
           REGION "GET ARRAY PARAMETERS"
               #len.tblData := UDINT_TO_DINT(CountOfElements(#tblData));
               #len.tblDisp := UDINT_TO_DINT(CountOfElements(#tblDisp));
           END_REGION

           REGION "CALCULATE UPPER BOUND"
               #ubound := #len.tblData;
               IF #first_null_index <= #len.tblData THEN
                   IF #first_null_index > 0 THEN
                       #ubound := #first_null_index;
                   END_IF;
               END_IF;
           END_REGION


           REGION "CALCULATE OFFSET"
               #offset := "Table Nav: Calculate Offset"(pulses := #pulses,
                                                        lenTblData := #ubound,
                                                        lenTblDisp := #len.tblDisp,
                                                        r1 := #r1);
           END_REGION


           REGION "CALCULATE FIRST ROW"
               #r1 := "Table Nav: Get First Row"(table_length := #ubound,
                                                 offset := #offset,
                                                 first_row := #r1);
           END_REGION


           REGION "CALCUALTE ROW INDICIES"
               "Table Nav: Calc Row Indices"(lenTblData := #ubound,
                                             lenTblDisp := #len.tblDisp,
                                             r1 := #r1,
                                             rowIndicies := #ret_row_indices);
           END_REGION


           REGION "RETURN ROW INDICIES"
               #RET_VAL := MOVE_BLK_VARIANT(SRC := #ret_row_indices,
                                            COUNT := DINT_TO_UDINT(#len.tblDisp),
                                            SRC_INDEX := 0,
                                            DEST_INDEX := 0,
                                            DEST => #rowIndices);
           END_REGION

       END_IF;
   END_REGION
END_FUNCTION_BLOCK

FUNCTION_BLOCK "Table Nav: Pulses"   // FB44, SCL
{ S7_Optimized_Access := 'TRUE' }
VERSION : 0.1
   VAR_INPUT
      press : "Nav Bar Data: PLC";
   END_VAR
   VAR_OUTPUT
      pulses : "Nav Bar Data: PLC";
   END_VAR
   VAR
      old : "Nav Bar Data: PLC";
   END_VAR
BEGIN
   REGION "EVALUATION"
       #pulses.top.actuate := #press.top.actuate AND NOT #old.top.actuate;
       #pulses.pageUp.actuate := #press.pageUp.actuate AND NOT #old.pageUp.actuate;
       #pulses.lineUp.actuate := #press.lineUp.actuate AND NOT #old.lineUp.actuate;
       #pulses.lineDown.actuate := #press.lineDown.actuate AND NOT #old.lineDown.actuate;
       #pulses.pageDown.actuate := #press.pageDown.actuate AND NOT #old.pageDown.actuate;
       #pulses.bottom.actuate := #press.bottom.actuate AND NOT #old.bottom.actuate;
   END_REGION

   REGION "CHANGE DETECTION"
       #old.top.actuate := #press.top.actuate;
       #old.pageUp.actuate := #press.pageUp.actuate;
       #old.lineUp.actuate := #press.lineUp.actuate;
       #old.lineDown.actuate := #press.lineDown.actuate;
       #old.pageDown.actuate := #press.pageDown.actuate;
       #old.bottom.actuate := #press.bottom.actuate;
   END_REGION
END_FUNCTION_BLOCK

FUNCTION "Table Nav: Get Null Index" : DInt   // FC14, SCL
{ S7_Optimized_Access := 'TRUE' }
VERSION : 0.1
   VAR_INPUT
      nullFlag : Int;
      nullCheckVals : Array[0.."WIP_COUNT"] of DInt;
   END_VAR
   VAR_TEMP
      pNullCheck : DInt;
   END_VAR
BEGIN
   WHILE #nullCheckVals[#pNullCheck] <> #nullFlag AND #pNullCheck <= "WIP_COUNT" DO
       #pNullCheck += 1;
   END_WHILE;
   #"Table Nav: Get Null Index" := #pNullCheck;
END_FUNCTION

FUNCTION "Table Nav: Get First Row" : DInt   // FC44, SCL
{ S7_Optimized_Access := 'TRUE' }
VERSION : 0.1
   VAR_INPUT
      first_row : DInt;
      offset : DInt;
      table_length : DInt;
   END_VAR
   VAR_TEMP
      ret : DInt;
   END_VAR
BEGIN
   REGION "DESCRIPTION"
       (*
       The new first row of the table is calculated from the offset. 
       Rollover and rollunder are resolved for the first row.
       *)
   END_REGION

   REGION "COPY TO INTERNAL"
       #ret := #first_row + #offset;
   END_REGION

   REGION "ROLLUNDER"
       IF #ret < 0 THEN
           #ret := #ret + #table_length;
       END_IF;
   END_REGION

   REGION "ROLLOVER"
       IF #ret > #table_length THEN
           #ret := #ret - #table_length;
       END_IF;
   END_REGION

   REGION "OUTPUT"
       #"Table Nav: Get First Row" := #ret;
   END_REGION
END_FUNCTION

FUNCTION "Table Nav: Calculate Offset" : DInt   // FC45, SCL
{ S7_Optimized_Access := 'TRUE' }
VERSION : 0.1
   VAR_INPUT
      lenTblData : DInt;
      lenTblDisp : DInt;
      pulses : "Nav Bar Data: PLC";
      r1 : DInt;
   END_VAR
   VAR_TEMP
      retOffset : DInt;
   END_VAR
   // Ret_Val : offset from table row 1 from button
BEGIN
   REGION "DESCRIPTION"
       (*
       The offset from the first row of the table is calculated based on the button pressed.
       *)
   END_REGION

   REGION "TOP"
       IF #pulses.top.actuate THEN
           #retOffset := -1 * #r1;
       END_IF;
   END_REGION

   REGION "PAGE UP"
       IF #pulses.pageUp.actuate THEN
           #retOffset := -1 * #lenTblDisp;
       END_IF;
   END_REGION

   REGION "LINE UP"
       IF #pulses.lineUp.actuate THEN
           #retOffset := -1;
       END_IF;
   END_REGION

   REGION "LINE DOWN"
       IF #pulses.lineDown.actuate THEN
           #retOffset := 1;
       END_IF;
   END_REGION

   REGION "PAGE DOWN"
       IF #pulses.pageDown.actuate THEN
           #retOffset := #lenTblDisp ;
       END_IF;
   END_REGION

   REGION "BOTTOM"
       IF #pulses.bottom.actuate THEN
           #retOffset := #lenTblData - #lenTblDisp - #r1;
       END_IF;
   END_REGION

   REGION "RETURN"
       #"Table Nav: Calculate Offset" := #retOffset;
   END_REGION
END_FUNCTION

FUNCTION "Table Nav: Calc Row Indices" : Void   // FC46, SCL
{ S7_Optimized_Access := 'TRUE' }
VERSION : 0.1
   VAR_INPUT
      lenTblData : DInt;
      lenTblDisp : DInt;
      r1 : DInt;
   END_VAR
   VAR_IN_OUT
      rowIndicies : Array[0..#lenRetArr] of DInt;
   END_VAR
   VAR_TEMP
      pOutArr : Int;
      calcRowIdx : DInt;
      retRowIndicies : Array[0..#lenRetArr] of DInt;
   END_VAR
   VAR CONSTANT
      lenRetArr : Int := 999;
   END_VAR
BEGIN
   REGION "DESCRIPTION"
       (*
       An array of the row indicies that the table should display is returned.
       Rollover and rollunder are calculated index by index.
       *) 
   END_REGION

   REGION "INITIALIZE OUTPUT"
       FOR #pOutArr := 0 TO #lenRetArr DO
           #rowIndicies[#pOutArr] := 0;
       END_FOR;
   END_REGION

   REGION "CALCULATE INDICIES"
       FOR #pOutArr := 0 TO DINT_TO_INT(#lenTblDisp) DO

           REGION "CALCULATE INDEX"
               #calcRowIdx := #r1 + INT_TO_DINT(#pOutArr);
           END_REGION

           REGION "ROLL UNDER"
               IF #calcRowIdx < 0 THEN
                   #calcRowIdx := #calcRowIdx + #lenTblDisp;
               END_IF;
           END_REGION

           REGION "ROLL OVER"
               IF #calcRowIdx >= #lenTblData THEN
                   #calcRowIdx := #calcRowIdx - #lenTblData;
               END_IF;
           END_REGION

           REGION "SAVE TO ARRAY"
               #retRowIndicies[#pOutArr] := #calcRowIdx;
           END_REGION

       END_FOR;
   END_REGION

   REGION "OUTPUT"
       #rowIndicies := #retRowIndicies;
   END_REGION
END_FUNCTION

FUNCTION "Table Nav: Run Trigger" : Bool   // FC47, SCL
{ S7_Optimized_Access := 'TRUE' }
VERSION : 0.1
   VAR_INPUT
      pulses : "Nav Bar Data: PLC";
   END_VAR
BEGIN
   #"Table Nav: Run Trigger" :=
       #pulses.top.actuate OR
       #pulses.pageUp.actuate OR
       #pulses.lineUp.actuate OR
       #pulses.lineDown.actuate OR
       #pulses.pageDown.actuate OR
       #pulses.bottom.actuate;
END_FUNCTION

// folder: Utilities/Time

FUNCTION "Time.to_WString" : WString   // FC36, SCL
{ S7_Optimized_Access := 'TRUE' }
VERSION : 0.1
   VAR_INPUT
      "Time" : Time;
   END_VAR
   VAR_TEMP
      _time : DInt;
      _days : DInt;
      _hours : DInt;
      _minutes : DInt;
      _seconds : DInt;
      "Time Elements" : Array[0..4] of WString;
      Length : Int;
      _return : WString;
   END_VAR
   VAR CONSTANT
      COLON : WString := WSTRING#':';
   END_VAR
BEGIN
   REGION GET INPUT
       #_time := #Time;
   END_REGION


   REGION CONVERT TIME INTO INDIVIDUAL PLACE VALUES
       #_days := "Time.Get_Days"(#_time);
       #_hours := "Time.Get_MOD_Hours"(#_time);
       #_minutes := "Time.Get_MOD_Minutes"(#_time);
       #_seconds := "Time.Get_MOD_Seconds"(#_time);
   END_REGION


   REGION "ASSEMBLE DISPLAY STRING"
       IF #_days > 0 THEN
           #_return := CONCAT_WSTRING(IN1 := #_return, IN2 := "Time.to_WString.Days"(#_time), IN3 := #COLON);
           #_return := CONCAT_WSTRING(IN1 := #_return, IN2 := "Time.to_WString.MOD_Hours"(#_time), IN3 := #COLON);
           #_return := CONCAT_WSTRING(IN1 := #_return, IN2 := "Time.to_WString.MOD_Minutes"(#_time), IN3 := #COLON);
           #_return := CONCAT_WSTRING(IN1 := #_return, IN2 := "Time.to_WString.MOD_Seconds"(#_time));
           #"Time.to_WString" := #_return;
           RETURN;
       END_IF;
       IF #_hours > 0 THEN
           #_return := CONCAT_WSTRING(IN1 := #_return, IN2 := "Time.to_WString.MOD_Hours"(#_time), IN3 := #COLON);
           #_return := CONCAT_WSTRING(IN1 := #_return, IN2 := "Time.to_WString.MOD_Minutes"(#_time), IN3 := #COLON);
           #_return := CONCAT_WSTRING(IN1 := #_return, IN2 := "Time.to_WString.MOD_Seconds"(#_time));
           #"Time.to_WString" := #_return;
           RETURN;
       END_IF;
       IF #_minutes > 0 THEN
           #_return := CONCAT_WSTRING(IN1 := #_return, IN2 := "Time.to_WString.MOD_Minutes"(#_time), IN3 := #COLON);
           #_return := CONCAT_WSTRING(IN1 := #_return, IN2 := "Time.to_WString.MOD_Seconds"(#_time));
           #"Time.to_WString" := #_return;
           RETURN;
       END_IF;
       IF #_seconds > 0 THEN
           #_return := CONCAT_WSTRING(IN1 := #_return, IN2 := "Time.to_WString.MOD_Seconds"(#_time));
           #"Time.to_WString" := #_return;
           RETURN;
       END_IF;
       #_return := WSTRING#'00:00';
       #"Time.to_WString" := #_return;
       RETURN;
   END_REGION
END_FUNCTION

FUNCTION "Time.to_WString.Seconds" : WString   // FC275, SCL
{ S7_Optimized_Access := 'TRUE' }
VERSION : 0.1
   VAR_INPUT
      value : Time;
   END_VAR
BEGIN
   #"Time.to_WString.Seconds" := "Time.to_WString.Prepare_Component"("Time.Get_Seconds"(#value));
END_FUNCTION

FUNCTION "Time.Get_MOD_Seconds" : DInt   // FC276, SCL
{ S7_Optimized_Access := 'TRUE' }
VERSION : 0.1
   VAR_INPUT
      value : Time;
   END_VAR
   VAR CONSTANT
      SECONDS_PER_MINUTE : DInt := 60;
   END_VAR
BEGIN
   #"Time.Get_MOD_Seconds" := "Time.Get_Seconds"(#value) MOD #SECONDS_PER_MINUTE;
END_FUNCTION

FUNCTION "Time.Get_MOD_Minutes" : DInt   // FC277, SCL
{ S7_Optimized_Access := 'TRUE' }
VERSION : 0.1
   VAR_INPUT
      value : Time;
   END_VAR
   VAR CONSTANT
      MINUTES_PER_HOUR : DInt := 60;
   END_VAR
BEGIN
   #"Time.Get_MOD_Minutes" := "Time.Get_Minutes"(#value) MOD #MINUTES_PER_HOUR;
END_FUNCTION

FUNCTION "Time.Get_MOD_Hours" : DInt   // FC278, SCL
{ S7_Optimized_Access := 'TRUE' }
VERSION : 0.1
   VAR_INPUT
      value : Time;
   END_VAR
   VAR CONSTANT
      HOURS_PER_DAY : DInt := 24;
   END_VAR
BEGIN
   #"Time.Get_MOD_Hours" := "Time.Get_Hours"(#value) MOD #HOURS_PER_DAY;
END_FUNCTION

FUNCTION "Time.Get_Days" : Int   // FC279, SCL
{ S7_Optimized_Access := 'TRUE' }
VERSION : 0.1
   VAR_INPUT
      value : Time;
   END_VAR
   VAR_TEMP
      _return : DInt;
   END_VAR
   VAR CONSTANT
      MILLISECONDS_PER_DAY : DInt := 86_000_000;
   END_VAR
BEGIN
   #_return := #value / #MILLISECONDS_PER_DAY;
   #"Time.Get_Days" := DINT_TO_INT(#_return);
END_FUNCTION

FUNCTION "Time.Get_Seconds" : DInt   // FC280, SCL
{ S7_Optimized_Access := 'TRUE' }
VERSION : 0.1
   VAR_INPUT
      value : Time;
   END_VAR
   VAR CONSTANT
      MILLISECONDS_PER_SECOND : DInt := 1_000;
   END_VAR
BEGIN
   #"Time.Get_Seconds" := #value / #MILLISECONDS_PER_SECOND;
END_FUNCTION

FUNCTION "Time.Get_Minutes" : DInt   // FC281, SCL
{ S7_Optimized_Access := 'TRUE' }
VERSION : 0.1
   VAR_INPUT
      value : Time;
   END_VAR
   VAR CONSTANT
      MILLISECONDS_PER_MINUTE : DInt := 60_000;
   END_VAR
BEGIN
   #"Time.Get_Minutes" := #value / #MILLISECONDS_PER_MINUTE;
END_FUNCTION

FUNCTION "Time.to_WString.Prepare_Component" : WString   // FC282, SCL
{ S7_Optimized_Access := 'TRUE' }
VERSION : 0.1
   VAR_INPUT
      component : DInt;
   END_VAR
   VAR_TEMP
      _return : WString;
   END_VAR
   VAR CONSTANT
      ZERO : WChar := WCHAR#'0';
   END_VAR
BEGIN
   #_return := DINT_TO_WSTRING(#component);
   #_return := "Trim"("Strip Sign"(#_return));
   #_return := "Add Leading"("Leading Character" := #ZERO,
                             "Desired Length" := 2,
                             "String" := #_return);
   #"Time.to_WString.Prepare_Component" := #_return;
END_FUNCTION

FUNCTION "Time.to_WString.Minutes" : WString   // FC284, SCL
{ S7_Optimized_Access := 'TRUE' }
VERSION : 0.1
   VAR_INPUT
      value : Time;
   END_VAR
   VAR_TEMP
      _to_udint : UDInt;
      _return : WString;
   END_VAR
BEGIN
   #"Time.to_WString.Minutes" := "Time.to_WString.Prepare_Component"("Time.Get_Minutes"(#value));
END_FUNCTION

FUNCTION "Time.to_WString.MOD_Minutes" : WString   // FC285, SCL
{ S7_Optimized_Access := 'TRUE' }
VERSION : 0.1
   VAR_INPUT
      value : Time;
   END_VAR
BEGIN
   #"Time.to_WString.MOD_Minutes" := "Time.to_WString.Prepare_Component"("Time.Get_MOD_Minutes"(#value));
END_FUNCTION

FUNCTION "Time.to_WString.Hours" : WString   // FC286, SCL
{ S7_Optimized_Access := 'TRUE' }
VERSION : 0.1
   VAR_INPUT
      value : Time;
   END_VAR
BEGIN
   #"Time.to_WString.Hours" := "Time.to_WString.Prepare_Component"("Time.Get_Hours"(#value));
END_FUNCTION

FUNCTION "Time.to_WString.MOD_Seconds" : WString   // FC287, SCL
{ S7_Optimized_Access := 'TRUE' }
VERSION : 0.1
   VAR_INPUT
      value : Time;
   END_VAR
BEGIN
   #"Time.to_WString.MOD_Seconds" := "Time.to_WString.Prepare_Component"("Time.Get_MOD_Seconds"(#value));
END_FUNCTION

FUNCTION "Time.Get_Hours" : DInt   // FC288, SCL
{ S7_Optimized_Access := 'TRUE' }
VERSION : 0.1
   VAR_INPUT
      value : Time;
   END_VAR
   VAR CONSTANT
      MILLISECONDS_PER_HOUR : DInt := 3_600_000;
   END_VAR
BEGIN
   #"Time.Get_Hours" := #value / #MILLISECONDS_PER_HOUR;
END_FUNCTION

FUNCTION "Time.to_WString.MOD_Hours" : WString   // FC290, SCL
{ S7_Optimized_Access := 'TRUE' }
VERSION : 0.1
   VAR_INPUT
      value : Time;
   END_VAR
BEGIN
   #"Time.to_WString.MOD_Hours" := "Time.to_WString.Prepare_Component"("Time.Get_MOD_Hours"(#value));
END_FUNCTION

FUNCTION "Time.to_WString.Days" : WString   // FC291, SCL
{ S7_Optimized_Access := 'TRUE' }
VERSION : 0.1
   VAR_INPUT
      value : Time;
   END_VAR
BEGIN
   #"Time.to_WString.Days" := "Time.to_WString.Prepare_Component"("Time.Get_Days"(#value));
END_FUNCTION

// folder: Utilities/Timer

FUNCTION "Timer.WString_to_Real" : Real   // FC39, SCL
{ S7_Optimized_Access := 'TRUE' }
VERSION : 0.1
   VAR_INPUT
      wstring : WString;
   END_VAR
   VAR CONSTANT
      msPerSec : Real := 1000.0;
   END_VAR
BEGIN
   #"Timer.WString_to_Real" := DINT_TO_REAL(TIME_TO_DINT("WString.to_Time"(#wstring))) / #msPerSec;
END_FUNCTION

FUNCTION "Timer.Real_to_WString" : WString   // FC40, SCL
{ S7_Optimized_Access := 'TRUE' }
VERSION : 0.1
   VAR_INPUT
      realVal : Real;
   END_VAR
   VAR CONSTANT
      msPerSec : Real := 1000.0;
   END_VAR
BEGIN
   #"Timer.Real_to_WString" := "Time.to_WString"(DINT_TO_TIME(REAL_TO_DINT(#realVal * #msPerSec)));
END_FUNCTION

FUNCTION "Timer" : Void   // FC79, SCL
{ S7_Optimized_Access := 'TRUE' }
VERSION : 0.1
   VAR_INPUT
      delta : Real;
      allotted : Real;
   END_VAR
   VAR_IN_OUT
      elapsed : Real;
      remaining : Real;
   END_VAR
   VAR_TEMP
      _elapsed : Real;
      _remaining : Real;
   END_VAR
BEGIN
   #_elapsed := #elapsed + #delta;
   #_remaining := #allotted - #_elapsed;
   #elapsed := #_elapsed;
   #remaining := #_remaining;
END_FUNCTION

FUNCTION "Timer.Digits_as_String_to_Seconds" : Time   // FC265, SCL
{ S7_Optimized_Access := 'TRUE' }
VERSION : 0.1
   VAR_INPUT
      digits : String;
   END_VAR
   VAR_TEMP
      _characters : Array[0..#CHAR_COUNT] of Char;
      _count : DInt;
      _i : Int;
      _length : Int;
      _character_count : Int;
      _return : DInt;
      _temp : Bool;
   END_VAR
   VAR CONSTANT
      ASCII_OFFSET : DInt := 16#30;
      BLANK : Time;
      CHAR_COUNT : Int := 9;
      MS_PER_SEC : DInt := 1_000;
   END_VAR
BEGIN
   REGION "EXIT ON NO INPUT"
       IF #digits = '' THEN
           #"Timer.Digits_as_String_to_Seconds" := #BLANK;
           RETURN;
       END_IF;
   END_REGION


   REGION "EXPLODE"
       Strg_TO_Chars(Strg := #digits,
                     pChars := 0,
                     Cnt => #_count,
                     Chars := #_characters);
       #_length := UDINT_TO_INT("Array.Any.Length"(#_characters)) - 1;
   END_REGION


   REGION "COUNT"
       #_character_count := "Array.Char.Search"(array := #_characters, search_term := ' ') - 1;
   END_REGION


   REGION "VALIDATE"
       FOR #_i := 0 TO #_character_count DO
           IF NOT "Char.Is_Numeric"(#_characters[#_i]) THEN
               #"Timer.Digits_as_String_to_Seconds" := #BLANK;
               RETURN;
           END_IF;
       END_FOR;
   END_REGION


   #"Timer.Digits_as_String_to_Seconds" := STRING_TO_DINT(#digits) * #MS_PER_SEC;
END_FUNCTION

FUNCTION "Timer.Digits_as_String_to_Minutes" : Time   // FC267, SCL
{ S7_Optimized_Access := 'TRUE' }
VERSION : 0.1
   VAR_INPUT
      digits : String;
   END_VAR
   VAR CONSTANT
      SECONDS_PER_MINUTE : Int := 60;
   END_VAR
BEGIN
   #"Timer.Digits_as_String_to_Minutes" := #SECONDS_PER_MINUTE * TIME_TO_DINT("Timer.Digits_as_String_to_Seconds"(#digits));
END_FUNCTION

FUNCTION "Timer.Digits_as_String_to_Hours" : Time   // FC269, SCL
{ S7_Optimized_Access := 'TRUE' }
VERSION : 0.1
   VAR_INPUT
      digits : String;
   END_VAR
   VAR CONSTANT
      SECONDS_PER_HOUR : Int := 3_600;
   END_VAR
BEGIN
   #"Timer.Digits_as_String_to_Hours" := #SECONDS_PER_HOUR * TIME_TO_DINT("Timer.Digits_as_String_to_Seconds"(#digits));
END_FUNCTION

// folder: Utilities/UInt

FUNCTION "UInt.Value_Change" : Bool   // FC183, SCL
{ S7_Optimized_Access := 'TRUE' }
VERSION : 0.1
   VAR_INPUT
      value : UInt;
      old_value : UInt;
   END_VAR
BEGIN
   #"UInt.Value_Change" := #value <> #old_value;
END_FUNCTION

// folder: Utilities/USInt

FUNCTION_BLOCK "USInt.State_change"   // FB58, SCL
{ S7_Optimized_Access := 'TRUE' }
VERSION : 0.1
   VAR_INPUT
      value : USInt;
   END_VAR
   VAR_IN_OUT
      get_usint : "State Changes: USInt";
   END_VAR
   VAR
      old_value : USInt;
   END_VAR
   VAR_TEMP
      _return : "State Changes: USInt";
   END_VAR
BEGIN
   REGION "BUFFER IN"
       #_return := #get_usint;
   END_REGION


   REGION "MAP"
       IF #value <> #old_value THEN
           #_return.actual := #value;
       END_IF;
       #_return.rising := "USInt.Rising_Edge"(value := #value,
                                              old_value := #old_value);
       #_return.falling := "USInt.Falling_Edge"(value := #value,
                                                old_value := #old_value);
   END_REGION


   REGION "SAVE OLD VALUE"
       #old_value := #_return.actual;
   END_REGION


   REGION "RETURN" 
       #get_usint := #_return;
   END_REGION
END_FUNCTION_BLOCK

FUNCTION "USInt.Value_Change" : Bool   // FC181, SCL
{ S7_Optimized_Access := 'TRUE' }
VERSION : 0.1
   VAR_INPUT
      value : USInt;
      old_value : USInt;
   END_VAR
BEGIN
   #"USInt.Value_Change" := #value <> #old_value;
END_FUNCTION

FUNCTION "USInt.Rising_Edge" : Bool   // FC262, SCL
{ S7_Optimized_Access := 'TRUE' }
VERSION : 0.1
   VAR_INPUT
      value : USInt;
      old_value : USInt;
   END_VAR
BEGIN
   #"USInt.Rising_Edge" := #value <> "NULL_TOKEN" AND #old_value = "NULL_TOKEN";
END_FUNCTION

FUNCTION "USInt.Falling_Edge" : Bool   // FC263, SCL
{ S7_Optimized_Access := 'TRUE' }
VERSION : 0.1
   VAR_INPUT
      value : USInt;
      old_value : USInt;
   END_VAR
BEGIN
   #"USInt.Falling_Edge" := #value = "NULL_TOKEN" AND #old_value <> "NULL_TOKEN";
END_FUNCTION

// folder: Utilities/WIP

FUNCTION "WIP.Code_to_WString" : WString   // FC64, SCL
{ S7_Optimized_Access := 'TRUE' }
VERSION : 0.1
   VAR_INPUT
      wipTxtLib : "Recipe: Wip Text Library";
      code : DInt;
   END_VAR
   VAR_TEMP
      wipCode : DInt;
      wipText : DInt;
      output : WString;
   END_VAR
   VAR CONSTANT
      newLine : WString := WSTRING#'$L';
   END_VAR
BEGIN
   REGION "PARSE CODE"
       "Part_Number.Parse_Code"(code := #code,
                    code_left => #wipCode,
                    code_right => #wipText);
   END_REGION

   REGION "DOUBLE LINE PN"
       #output := CONCAT_WSTRING(IN1 := #wipTxtLib.code[#wipCode],
                                 IN2 := #newLine,
                                 IN3 := #wipTxtLib.txt[#wipText]);
   END_REGION

   REGION "OUTPUT"
       #"WIP.Code_to_WString" := #output;
   END_REGION
END_FUNCTION

FUNCTION "WIP.Count" : Int   // FC72, SCL
{ S7_Optimized_Access := 'TRUE' }
VERSION : 0.1
   VAR_INPUT
      stnSavedWips : "WIP: Station";
   END_VAR
   VAR_TEMP
      pWip : Int;
   END_VAR
   // Ret_Val : -1 for no wips in station
BEGIN
   WHILE #stnSavedWips.wip[#pWip].wip.code <> -1 DO
       #pWip += 1;
   END_WHILE;
   #"WIP.Count" := #pWip - 1;
END_FUNCTION

FUNCTION "WIP.Global_Index_to_Station" : "WIP: Station"   // FC113, SCL
{ S7_Optimized_Access := 'TRUE' }
VERSION : 0.1
   VAR_INPUT
      index : Int;
      wip_stations : "Recipe: HMI Stations Saved Wips";
   END_VAR
   VAR_TEMP
      i : Int;
      ret : "WIP: Station";
   END_VAR
BEGIN
   REGION "FIND STATION"
       FOR #i := 0 TO "HMI_STATION_COUNT" DO
           IF #wip_stations.stn[#i].pStn = #index THEN
               #ret := #wip_stations.stn[#i];
               EXIT;
           END_IF;
       END_FOR;
   END_REGION


   REGION "RETURN"
       #"WIP.Global_Index_to_Station" := #ret;
   END_REGION
END_FUNCTION

FUNCTION "WIP.Global_Index_to_HMI_Station_Index" : Int   // FC130, SCL
{ S7_Optimized_Access := 'TRUE' }
VERSION : 0.1
   VAR_INPUT
      global_index : Int;
      saved_WIPs : "Recipe: HMI Stations Saved Wips";
   END_VAR
   VAR_TEMP
      i : Int;
      ret : Int;
   END_VAR
BEGIN
   REGION "SEARCH FOR INDEX"
       #ret := "NULL_TOKEN";
       FOR #i := 0 TO "HMI_STATION_COUNT" DO
           IF #saved_WIPs.stn[#i].pStn = #global_index THEN
               #ret := #i;
               EXIT;
           END_IF;
       END_FOR;
   END_REGION


   REGION "RETURN"
       #"WIP.Global_Index_to_HMI_Station_Index" := #ret;
   END_REGION
END_FUNCTION

FUNCTION "WIP.Code_to_Index" : Int   // FC233, SCL
{ S7_Optimized_Access := 'TRUE' }
VERSION : 0.1
   VAR_INPUT
      saved_wip : "WIP: Station";
      wip_code : DInt;
   END_VAR
   VAR_TEMP
      _i : Int;
      _length : Int;
   END_VAR
BEGIN
   #_length := UDINT_TO_INT("Array.Any.Length"(#saved_wip.wip)) - 1;
   FOR #_i := 0 TO #_length DO
       IF #wip_code <> #saved_wip.wip[#_i].wip.code THEN
           CONTINUE;
       END_IF;
       #"WIP.Code_to_Index" := #_i;
       RETURN;
   END_FOR;

   #"WIP.Code_to_Index" := "NULL_TOKEN";
   RETURN;
END_FUNCTION

FUNCTION "WIP_Station.Indices_of_Selected_WIPs" : Void   // FC241, SCL
{ S7_Optimized_Access := 'TRUE' }
VERSION : 0.1
   VAR_INPUT
      selected_wips : "Selected Wips";
      station_wips : "WIP: Station";
   END_VAR
   VAR_IN_OUT
      selected_wip_indices : Array[*] of Int;
   END_VAR
   VAR_TEMP
      _i : Int;
      _length : Int;
      _p_return : Int;
      _wip_index : Int;
   END_VAR
   VAR CONSTANT
      UBOUND : Int := 999;
   END_VAR
BEGIN
   REGION "PREP ARRAY OF FOUND INDICES"
       "Array.Int.Fill"(value := "NULL_TOKEN",
                        int_array := #selected_wip_indices);
       #_length := UDINT_TO_INT("Array.Any.Length"(#selected_wip_indices)) - 1;
   END_REGION

   REGION "FOR EACH SELECTED WIP"
       FOR #_i := 0 TO #selected_wips.count - 1 DO

           REGION "GET SELECTED WIPS INDEX IN THIS STATION"
               #_wip_index := "WIP_Station.Indices_of_Selected_WIPS.Search_WIP"(wip_code := #selected_wips.wips[#_i],
                                                                                station_wips := #station_wips);
           END_REGION

           REGION "IF NOT FOUND GO TO NEXT WIP"
               // fault tolerance
               IF #_wip_index = "NULL_TOKEN" THEN
                   CONTINUE;
               END_IF;
           END_REGION

           REGION "WIP FOUND IN STATION"
               #selected_wip_indices[#_p_return] := #_wip_index;
               #_p_return += 1;
           END_REGION

           REGION "DON'T GO OUT OF FOUND IDEX ARRAY"
               // fault tolerance
               IF #_p_return > #_length THEN
                   RETURN;
               END_IF;
           END_REGION

       END_FOR;
   END_REGION
END_FUNCTION

FUNCTION "WIP_Station.Indices_of_Selected_WIPS.Search_WIP" : Int   // FC242, SCL
{ S7_Optimized_Access := 'TRUE' }
VERSION : 0.1
   VAR_INPUT
      wip_code : DInt;
      station_wips : "WIP: Station";
   END_VAR
   VAR_TEMP
      _i : Int;
      _length : Int;
   END_VAR
BEGIN
   REGION "FOR EACH WIP IN STATION"
       #_length := UDINT_TO_INT("Array.Any.Length"(#station_wips.wip)) - 1;
       FOR #_i := 0 TO #_length DO

           REGION "WIP CODE DOES NOT MATCH"
               IF #wip_code <> #station_wips.wip[#_i].wip.code THEN
                   CONTINUE;
               END_IF;
           END_REGION

           REGION "WIP CODE MATCHES"
               #"WIP_Station.Indices_of_Selected_WIPS.Search_WIP" := #_i;
               RETURN;
           END_REGION

       END_FOR;
   END_REGION

   REGION "NO MATCH FOUND"
       #"WIP_Station.Indices_of_Selected_WIPS.Search_WIP" := "NULL_TOKEN";
       RETURN;
   END_REGION
END_FUNCTION

// folder: Utilities/WString

FUNCTION_BLOCK "WString.State_Change"   // FB51, SCL
{ S7_Optimized_Access := 'TRUE' }
VERSION : 0.1
   VAR_INPUT
      interface : WString;
   END_VAR
   VAR_IN_OUT
      get_wstring : "State Changes: WString";
   END_VAR
   VAR
      old_value : WString;
   END_VAR
   VAR_TEMP
      ret : "State Changes: WString";
   END_VAR
   VAR CONSTANT
      blank : WString;
   END_VAR
BEGIN
   REGION "BUFFER IN"
       #ret := #get_wstring;
   END_REGION


   REGION "MAP"
       IF #interface <> #old_value THEN
           #ret.actual := #interface;
       END_IF;
       #ret.rising := "WString.Rising_Edge"(value := #interface,
                                             old_value := #old_value);
       #ret.falling := "WString.Falling_Edge"(value := #interface,
                                               old_value := #old_value);
   END_REGION


   REGION "SAVE OLD VALUE"
       #old_value := #ret.actual;
   END_REGION


   REGION "RETURN" 
       #get_wstring := #ret;
   END_REGION
END_FUNCTION_BLOCK

FUNCTION "WString.to_Time" : Time   // FC38, SCL
{ S7_Optimized_Access := 'TRUE' }
VERSION : 0.1
   VAR_INPUT
      value : WString;
   END_VAR
   VAR_TEMP
      _component_count : Int;
      _i : Int;
      _return : DInt;
      _time_components : Array[0..4] of WString;
   END_VAR
   VAR CONSTANT
      BLANK : Time;
   END_VAR
BEGIN
   REGION "NO INPUT"
       IF #value = WSTRING#'' THEN
           #"WString.to_Time" := #BLANK;
           RETURN;
       END_IF;
   END_REGION


   REGION "NO DELIMETERS"
       IF FIND(IN1 := WSTRING_TO_STRING(#value), IN2 := ':') = 0 THEN
           IF NOT "WString.to_Time.Validate_Component"(WSTRING_TO_STRING(#value)) THEN
               #"WString.to_Time" := #BLANK;
               RETURN;
           END_IF;
           #_return := "Timer.Digits_as_String_to_Seconds"(WSTRING_TO_STRING(#value));
       END_IF;
   END_REGION


   REGION "EXPLODE INPUT"
       "WString.Split_Single"(wstring_in := #value,
                              delimeter := WString#':',
                              "pointer" := 0,
                              sub_strings := #_time_components);
       #_component_count := "Array.WString.Search"(array := #_time_components, search_term := WString#'') - 1;
   END_REGION


   REGION "EXIT ON TOO MANY COMPONENTS"
       IF #_component_count >= 3 THEN
           #"WString.to_Time" := #BLANK;
       END_IF;
   END_REGION


   REGION "VALIDATE INPUT"
       FOR #_i := 0 TO #_component_count DO
           IF NOT "WString.to_Time.Validate_Component"(WSTRING_TO_STRING(#_time_components[#_i])) THEN
               #"WString.to_Time" := #BLANK;
               RETURN;
           END_IF;
       END_FOR;
   END_REGION


   REGION "REVERSE"
       "Array.WString.Reverse"(null_token := wstring#'',
                               wstring_array := #_time_components);
   END_REGION


   REGION CONVERT ARRAY ELEMENTS TO TIME
       #_return := 0;
       FOR #_i := 0 TO #_component_count DO
           CASE #_i OF
               0:
                   #_return := TIME_TO_DINT("Timer.Digits_as_String_to_Seconds"(WSTRING_TO_STRING(#_time_components[#_i])));
               1:
                   #_return += TIME_TO_DINT("Timer.Digits_as_String_to_Minutes"(WSTRING_TO_STRING(#_time_components[#_i])));
               2:
                   #_return += TIME_TO_DINT("Timer.Digits_as_String_to_Hours"(WSTRING_TO_STRING(#_time_components[#_i])));
           END_CASE;
       END_FOR;
   END_REGION


   REGION RETURN VALUE

       #"WString.to_Time" := DINT_TO_TIME(#_return);

   END_REGION
END_FUNCTION

FUNCTION "WString.Rising_Edge" : Bool   // FC182, SCL
{ S7_Optimized_Access := 'TRUE' }
VERSION : 0.1
   VAR_INPUT
      value : WString;
      old_value : WString;
   END_VAR
   VAR CONSTANT
      blank : WString;
   END_VAR
BEGIN
   #"WString.Rising_Edge" := #value <> #blank AND #old_value = #blank;
END_FUNCTION

FUNCTION "WString.Falling_Edge" : Bool   // FC188, SCL
{ S7_Optimized_Access := 'TRUE' }
VERSION : 0.1
   VAR_INPUT
      value : WString;
      old_value : WString;
   END_VAR
   VAR CONSTANT
      blank : WString;
   END_VAR
BEGIN
   #"WString.Falling_Edge" := #value = #blank AND #old_value <> #blank;
END_FUNCTION

FUNCTION "WString.to_Time.Validate_Component" : Bool   // FC273, SCL
{ S7_Optimized_Access := 'TRUE' }
VERSION : 0.1
   VAR_INPUT
      component : String;
   END_VAR
   VAR_TEMP
      _characters : Array[0..#CHAR_COUNT] of Char;
      _character_count : Int;
      _count : DInt;
      _i : Int;
   END_VAR
   VAR CONSTANT
      CHAR_COUNT : Int := 9;
   END_VAR
BEGIN
   Strg_TO_Chars(Strg := #component,
                 pChars := 0,
                 Cnt => #_count,
                 Chars := #_characters);
   #_character_count := "Array.Char.Search"(array := #_characters, search_term := ' ') - 1;
   FOR #_i := 0 TO #_character_count DO
       IF NOT "Char.Is_Numeric"(#_characters[#_i]) THEN
           #"WString.to_Time.Validate_Component" := FALSE;
           RETURN;
       END_IF;
   END_FOR;
   #"WString.to_Time.Validate_Component" := TRUE;
   RETURN;
END_FUNCTION

// ===== library types =====

TYPE "PB Data"
   STRUCT
      actuate : Bool;
      animate : USInt;
      enable : Bool;
      label : WString[80];
      listSelect : UInt;
      visible : Bool;
   END_STRUCT;
END_TYPE

TYPE "PB Data: Text Label"
   STRUCT
      actuate : Bool;
      animate : USInt;
      label : WString[20];
   END_STRUCT;
END_TYPE

TYPE "Station Assignment: Button Details Data"
   STRUCT
      alloted : Struct
         animate : USInt;
         value : WString[10];
      END_STRUCT;
      critical : Struct
         animate : USInt;
         value : WString[10];
      END_STRUCT;
      label : Struct
         animate : USInt;
         value : WString[2];
      END_STRUCT;
      partNumber : Struct
         animate : USInt;
         value : WString[40];
      END_STRUCT;
      select : Struct
         actuate : Bool;
         animate : USInt;
      END_STRUCT;
   END_STRUCT;
END_TYPE

TYPE "IO Field Data: Timers"
   STRUCT
      animate : USInt;
      inputFinished : Bool;
      value : WString[5];
   END_STRUCT;
END_TYPE

TYPE "Line Label Data"
   STRUCT
      animate : Struct
         bg : USInt;
         ioField : USInt;
      END_STRUCT;
      inputFinished : Bool;
      value : WString[10];
   END_STRUCT;
END_TYPE

TYPE "IO Field Data: Part Number: 2 Line"
   STRUCT
      single_actuate : Bool;
      single_animate : USInt;
      single_enable : Bool;
      single_input_finished : Bool;
      single_value : WString[40];
      single_visible : Bool;
      double_actuate : Bool;
      double_animate : USInt;
      double_enable : Bool;
      double_input_finished_top : Bool;
      double_input_finished_bottom : Bool;
      double_value_top : WString[40];
      double_value_bottom : WString[40];
      double_visible : Bool;
   END_STRUCT;
END_TYPE

TYPE "Drop Zone Data"
   STRUCT
      animate : Struct
         bg : USInt;
         ioField : USInt;
      END_STRUCT;
      inputFinished : Bool;
      value : WString[10];
   END_STRUCT;
END_TYPE

TYPE "Station Sim Data"
   STRUCT
      stn : Struct
         animate : USInt;
         label : WString[20];
      END_STRUCT;
      btn : Struct
         actuate : Byte;
         animate : Array[0..7] of USInt;
         labels : Array[0..7] of WString [4];
      END_STRUCT;
   END_STRUCT;
END_TYPE

// folder: Main HMI

TYPE "Table Row Data"
   STRUCT
      address : DInt := -1;
      ordered : Bool;
      pbSelection : Struct
         actuate : Bool;
         animate : USInt;
      END_STRUCT;
      rtBackground : Struct
         animate : USInt;
      END_STRUCT;
      tfDropZone : Struct
         animate : USInt;
         value : WString[20];
      END_STRUCT;
      tfLine : Struct
         animate : USInt;
         value : WString[20];
      END_STRUCT;
      tfPartNumber : Struct
         animateDL : USInt;
         animateSL : USInt;
         value : WString[40];
      END_STRUCT;
      tfTime : Struct
         animate : USInt;
         value : WString[20];
      END_STRUCT;
   END_STRUCT;
END_TYPE

(* ===== HMI "HMI_RT_1" =====
system functions are stored by id; their names below are inferred from use
connection "Main HMI": ETHERNET, S7_1500_OMS

HMI tags "Default tag table"
   "Clock_Byte" : Byte = PLC Clock_Byte AT %MB0, 100 ms
   "HMI Data: Warehouse HMI_screenNumber" : Int = PLC "HMI Data: Warehouse HMI".screenNumber AT %DB1.DBW0, 100 ms
   "HMI Data: Warehouse HMI_barcode" : Barcode.UDT = PLC "HMI Data: Warehouse HMI".barcode AT %DB1.DBW0, 100 ms
   "HMI Data: Warehouse HMI_tableNav_top" : Push Button Data = PLC "HMI Data: Warehouse HMI".tableNav.top, 100 ms
   "HMI Data: Warehouse HMI_tableNav_pageUp" : Push Button Data = PLC "HMI Data: Warehouse HMI".tableNav.pageUp, 100 ms
   "HMI Data: Warehouse HMI_tableNav_lineUp" : Push Button Data = PLC "HMI Data: Warehouse HMI".tableNav.lineUp, 100 ms
   "HMI Data: Warehouse HMI_tableNav_lineDown" : Push Button Data = PLC "HMI Data: Warehouse HMI".tableNav.lineDown, 100 ms
   "HMI Data: Warehouse HMI_tableNav_pageDown" : Push Button Data = PLC "HMI Data: Warehouse HMI".tableNav.pageDown, 100 ms
   "HMI Data: Warehouse HMI_tableNav_bottom" : Push Button Data = PLC "HMI Data: Warehouse HMI".tableNav.bottom, 100 ms
   "HMI Data: Warehouse HMI_networkHealth_pnioDevices{1}" : Push Button Data = PLC "HMI Data: Warehouse HMI".networkHealth.pnioDevices[1], 100 ms
   "HMI Data: Warehouse HMI_networkHealth_pnioDevices{2}" : Push Button Data = PLC "HMI Data: Warehouse HMI".networkHealth.pnioDevices[2], 100 ms
   "HMI Data: Warehouse HMI_networkHealth_pnioDevices{3}" : Push Button Data = PLC "HMI Data: Warehouse HMI".networkHealth.pnioDevices[3], 100 ms
   "HMI Data: Warehouse HMI_networkHealth_pnioDevices{4}" : Push Button Data = PLC "HMI Data: Warehouse HMI".networkHealth.pnioDevices[4], 100 ms
   "HMI Data: Warehouse HMI_networkHealth_pnioDevices{5}" : Push Button Data = PLC "HMI Data: Warehouse HMI".networkHealth.pnioDevices[5], 100 ms
   "HMI Data: Warehouse HMI_networkHealth_pnioDevices{6}" : Push Button Data = PLC "HMI Data: Warehouse HMI".networkHealth.pnioDevices[6], 100 ms
   "HMI Data: Warehouse HMI_networkHealth_pnioDevices{7}" : Push Button Data = PLC "HMI Data: Warehouse HMI".networkHealth.pnioDevices[7], 100 ms
   "HMI Data: Warehouse HMI_networkHealth_pnioDevices{8}" : Push Button Data = PLC "HMI Data: Warehouse HMI".networkHealth.pnioDevices[8], 100 ms
   "HMI Data: Warehouse HMI_networkHealth_pnioDevices{9}" : Push Button Data = PLC "HMI Data: Warehouse HMI".settings.selectStation, 100 ms
   "HMI Data: Warehouse HMI_networkHealth_pnioDevices{10}" : Push Button Data = PLC "HMI Data: Warehouse HMI".networkHealth.pnioDevices[10], 100 ms
   "HMI Data: Warehouse HMI_networkHealth_pnioDevices{11}" : Push Button Data = PLC "HMI Data: Warehouse HMI".networkHealth.pnioDevices[11], 100 ms
   "HMI Data: Warehouse HMI_networkHealth_pnioDevices{12}" : Push Button Data = PLC "HMI Data: Warehouse HMI".networkHealth.pnioDevices[12], 100 ms
   "HMI Data: Warehouse HMI_networkHealth_pnioDevices{13}" : Push Button Data = PLC "HMI Data: Warehouse HMI".networkHealth.pnioDevices[13], 100 ms
   "HMI Data: Warehouse HMI_networkHealth_pnioDevices{16}" : Push Button Data = PLC "HMI Data: Warehouse HMI".networkHealth.pnioDevices[16], 100 ms
   "HMI Data: Warehouse HMI_networkHealth_pnioDevices{14}" : Push Button Data = PLC "HMI Data: Warehouse HMI".networkHealth.pnioDevices[14], 100 ms
   "HMI Data: Warehouse HMI_networkHealth_pnioDevices{15}" : Push Button Data = PLC "HMI Data: Warehouse HMI".networkHealth.pnioDevices[15], 100 ms
   "HMI Data: Warehouse HMI_networkHealth_pnioDevices{17}" : Push Button Data = PLC "HMI Data: Warehouse HMI".networkHealth.pnioDevices[17], 100 ms
   "HMI Data: Warehouse HMI_networkHealth_pnioDevices{18}" : Push Button Data = PLC "HMI Data: Warehouse HMI".networkHealth.pnioDevices[18], 100 ms
   "HMI Data: Warehouse HMI_networkHealth_pnioDevices{19}" : Push Button Data = PLC "HMI Data: Warehouse HMI".networkHealth.pnioDevices[19], 100 ms
   "HMI Data: Warehouse HMI_networkHealth_pnioDevices{20}" : Push Button Data = PLC "HMI Data: Warehouse HMI".networkHealth.pnioDevices[20], 100 ms
   "HMI Data: Warehouse HMI_networkHealth_pnioDevices{21}" : Push Button Data = PLC "HMI Data: Warehouse HMI".networkHealth.pnioDevices[21], 100 ms
   "HMI Data: Warehouse HMI_networkHealth_pnioDevices{22}" : Push Button Data = PLC "HMI Data: Warehouse HMI".networkHealth.pnioDevices[22], 100 ms
   "HMI Data: Warehouse HMI_networkHealth_pnioDevices{31}" : Push Button Data = PLC "HMI Data: Warehouse HMI".networkHealth.pnioDevices[31], 100 ms
   "HMI Data: Warehouse HMI_networkHealth_pnioDevices{32}" : Push Button Data = PLC "HMI Data: Warehouse HMI".networkHealth.pnioDevices[32], 100 ms
   "HMI Data: Warehouse HMI_networkHealth_pnioDevices{29}" : Push Button Data = PLC "HMI Data: Warehouse HMI".networkHealth.pnioDevices[29], 100 ms
   "HMI Data: Warehouse HMI_networkHealth_pnioDevices{30}" : Push Button Data = PLC "HMI Data: Warehouse HMI".networkHealth.pnioDevices[30], 100 ms
   "HMI Data: Warehouse HMI_networkHealth_pnioDevices{27}" : Push Button Data = PLC "HMI Data: Warehouse HMI".networkHealth.pnioDevices[27], 100 ms
   "HMI Data: Warehouse HMI_networkHealth_pnioDevices{28}" : Push Button Data = PLC "HMI Data: Warehouse HMI".networkHealth.pnioDevices[28], 100 ms
   "HMI Data: Warehouse HMI_networkHealth_pnioDevices{23}" : Push Button Data = PLC "HMI Data: Warehouse HMI".networkHealth.pnioDevices[23], 100 ms
   "HMI Data: Warehouse HMI_networkHealth_pnioDevices{24}" : Push Button Data = PLC "HMI Data: Warehouse HMI".networkHealth.pnioDevices[24], 100 ms
   "HMI Data: Warehouse HMI_networkHealth_pnioDevices{25}" : Push Button Data = PLC "HMI Data: Warehouse HMI".networkHealth.pnioDevices[25], 100 ms
   "HMI Data: Warehouse HMI_networkHealth_pnioDevices{26}" : Push Button Data = PLC "HMI Data: Warehouse HMI".networkHealth.pnioDevices[26], 100 ms
   "HMI Data: Warehouse HMI_networkHealth_pnioDevices{33}" : Push Button Data = PLC "HMI Data: Warehouse HMI".networkHealth.pnioDevices[33], 100 ms
   "HMI Data: Warehouse HMI_networkHealth_pnioDevices{34}" : Push Button Data = PLC "HMI Data: Warehouse HMI".networkHealth.pnioDevices[34], 100 ms
   "HMI Data: Warehouse HMI_networkHealth_pnioDevices{35}" : Push Button Data = PLC "HMI Data: Warehouse HMI".networkHealth.pnioDevices[35], 100 ms
   "HMI Data: Warehouse HMI_networkHealth_pnioDevices{36}" : Push Button Data = PLC "HMI Data: Warehouse HMI".networkHealth.pnioDevices[36], 100 ms
   "HMI Data: Warehouse HMI_networkHealth_pnioDevices{37}" : Push Button Data = PLC "HMI Data: Warehouse HMI".networkHealth.pnioDevices[37], 100 ms
   "HMI Data: Warehouse HMI_networkHealth_pnioDevices{38}" : Push Button Data = PLC "HMI Data: Warehouse HMI".networkHealth.pnioDevices[38], 100 ms
   "HMI Data: Warehouse HMI_networkHealth_pnioDevices{39}" : Push Button Data = PLC "HMI Data: Warehouse HMI".networkHealth.pnioDevices[39], 100 ms
   "HMI Data: Warehouse HMI_networkHealth_pnioDevices{40}" : Push Button Data = PLC "HMI Data: Warehouse HMI".networkHealth.pnioDevices[40], 100 ms
   "HMI Data: Warehouse HMI_networkHealth_pnioDevices{41}" : Push Button Data = PLC "HMI Data: Warehouse HMI".networkHealth.pnioDevices[41], 100 ms
   "HMI Data: Warehouse HMI_networkHealth_pnioDevices{42}" : Push Button Data = PLC "HMI Data: Warehouse HMI".networkHealth.pnioDevices[42], 100 ms
   "HMI Data: Warehouse HMI_networkHealth_pnioDevices{43}" : Push Button Data = PLC "HMI Data: Warehouse HMI".networkHealth.pnioDevices[43], 100 ms
   "HMI Data: Warehouse HMI_networkHealth_pnioDevices{44}" : Push Button Data = PLC "HMI Data: Warehouse HMI".networkHealth.pnioDevices[44], 100 ms
   "HMI Data: Warehouse HMI_networkHealth_pnioDevices{45}" : Push Button Data = PLC "HMI Data: Warehouse HMI".networkHealth.pnioDevices[45], 100 ms
   "HMI Data: Warehouse HMI_networkHealth_pnioDevices{46}" : Push Button Data = PLC "HMI Data: Warehouse HMI".networkHealth.pnioDevices[46], 100 ms
   "HMI Data: Warehouse HMI_networkHealth_pnioDevices{47}" : Push Button Data = PLC "HMI Data: Warehouse HMI".networkHealth.pnioDevices[47], 100 ms
   "HMI Data: Warehouse HMI_networkHealth_pnioDevices{48}" : Push Button Data = PLC "HMI Data: Warehouse HMI".networkHealth.pnioDevices[48], 100 ms
   "HMI Data: Warehouse HMI_networkHealth_et200spPopUp" : Station: ET200SP Comm Debug Data = PLC "HMI Data: Warehouse HMI".networkHealth.et200spPopUp, 100 ms
   "HMI Data: Warehouse HMI_networkHealth_kp8PopUp" : Station: KP8 Comm Debug Data = PLC "HMI Data: Warehouse HMI".networkHealth.kp8PopUp, 100 ms
   "HMI Data: Warehouse HMI_networkHealth_selectedDevice" : Int = PLC "HMI Data: Warehouse HMI".networkHealth.selectedDevice, 100 ms

HMI tags "Pop Ups: Select Buttons"
   "HMI Data: Warehouse HMI_pop_up_select_buttons_buttons{0}" : Push Button Data = PLC "HMI Data: Warehouse HMI".pop_up.select_buttons.buttons[0], 100 ms
   "HMI Data: Warehouse HMI_pop_up_select_buttons_buttons{1}" : Push Button Data = PLC "HMI Data: Warehouse HMI".pop_up.select_buttons.buttons[1], 100 ms
   "HMI Data: Warehouse HMI_pop_up_select_buttons_buttons{2}" : Push Button Data = PLC "HMI Data: Warehouse HMI".pop_up.select_buttons.buttons[2], 100 ms
   "HMI Data: Warehouse HMI_pop_up_select_buttons_buttons{3}" : Push Button Data = PLC "HMI Data: Warehouse HMI".pop_up.select_buttons.buttons[3], 100 ms
   "HMI Data: Warehouse HMI_pop_up_select_buttons_buttons{4}" : Push Button Data = PLC "HMI Data: Warehouse HMI".pop_up.select_buttons.buttons[4], 100 ms
   "HMI Data: Warehouse HMI_pop_up_select_buttons_buttons{5}" : Push Button Data = PLC "HMI Data: Warehouse HMI".pop_up.select_buttons.buttons[5], 100 ms
   "HMI Data: Warehouse HMI_pop_up_select_buttons_buttons{6}" : Push Button Data = PLC "HMI Data: Warehouse HMI".pop_up.select_buttons.buttons[6], 100 ms
   "HMI Data: Warehouse HMI_pop_up_select_buttons_buttons{7}" : Push Button Data = PLC "HMI Data: Warehouse HMI".pop_up.select_buttons.buttons[7], 100 ms
   "HMI Data: Warehouse HMI_pop_up_select_buttons_close_screen" : Push Button Data = PLC "HMI Data: Warehouse HMI".pop_up.select_buttons.close_screen, 100 ms

HMI tags "Pop Ups: Select Stations"
   "HMI Data: Warehouse HMI_pop_up_select_stations_close_screen" : Push Button Data = PLC "HMI Data: Warehouse HMI".pop_up.select_stations.close_screen, 100 ms
   "HMI Data: Warehouse HMI_pop_up_select_stations_nav_bar_hmi" : Nav Bar Data: HMI = PLC "HMI Data: Warehouse HMI".pop_up.select_stations.nav_bar.hmi, 100 ms
   "HMI Data: Warehouse HMI_pop_up_select_stations_stn_select_btns{0}" : Push Button Data = PLC "HMI Data: Warehouse HMI".pop_up.select_stations.stn_select_btns[0], 100 ms
   "HMI Data: Warehouse HMI_pop_up_select_stations_stn_select_btns{1}" : Push Button Data = PLC "HMI Data: Warehouse HMI".pop_up.select_stations.stn_select_btns[1], 100 ms
   "HMI Data: Warehouse HMI_pop_up_select_stations_stn_select_btns{10}" : Push Button Data = PLC "HMI Data: Warehouse HMI".pop_up.select_stations.stn_select_btns[10], 100 ms
   "HMI Data: Warehouse HMI_pop_up_select_stations_stn_select_btns{11}" : Push Button Data = PLC "HMI Data: Warehouse HMI".pop_up.select_stations.stn_select_btns[11], 100 ms
   "HMI Data: Warehouse HMI_pop_up_select_stations_stn_select_btns{2}" : Push Button Data = PLC "HMI Data: Warehouse HMI".pop_up.select_stations.stn_select_btns[2], 100 ms
   "HMI Data: Warehouse HMI_pop_up_select_stations_stn_select_btns{3}" : Push Button Data = PLC "HMI Data: Warehouse HMI".pop_up.select_stations.stn_select_btns[3], 100 ms
   "HMI Data: Warehouse HMI_pop_up_select_stations_stn_select_btns{4}" : Push Button Data = PLC "HMI Data: Warehouse HMI".pop_up.select_stations.stn_select_btns[4], 100 ms
   "HMI Data: Warehouse HMI_pop_up_select_stations_stn_select_btns{5}" : Push Button Data = PLC "HMI Data: Warehouse HMI".pop_up.select_stations.stn_select_btns[5], 100 ms
   "HMI Data: Warehouse HMI_pop_up_select_stations_stn_select_btns{6}" : Push Button Data = PLC "HMI Data: Warehouse HMI".pop_up.select_stations.stn_select_btns[6], 100 ms
   "HMI Data: Warehouse HMI_pop_up_select_stations_stn_select_btns{7}" : Push Button Data = PLC "HMI Data: Warehouse HMI".pop_up.select_stations.stn_select_btns[7], 100 ms
   "HMI Data: Warehouse HMI_pop_up_select_stations_stn_select_btns{8}" : Push Button Data = PLC "HMI Data: Warehouse HMI".pop_up.select_stations.stn_select_btns[8], 100 ms
   "HMI Data: Warehouse HMI_pop_up_select_stations_stn_select_btns{9}" : Push Button Data = PLC "HMI Data: Warehouse HMI".pop_up.select_stations.stn_select_btns[9], 100 ms

HMI tags "Pop Ups: Select WIPs"
   "HMI Data: Warehouse HMI_pop_up_select_WIPs_select_wip_buttons{0}" : Push Button Data = PLC "HMI Data: Warehouse HMI".pop_up.select_WIPs.select_wip_buttons[0], 100 ms
   "HMI Data: Warehouse HMI_pop_up_select_WIPs_select_wip_buttons{1}" : Push Button Data = PLC "HMI Data: Warehouse HMI".pop_up.select_WIPs.select_wip_buttons[1], 100 ms
   "HMI Data: Warehouse HMI_pop_up_select_WIPs_select_wip_buttons{2}" : Push Button Data = PLC "HMI Data: Warehouse HMI".pop_up.select_WIPs.select_wip_buttons[2], 100 ms
   "HMI Data: Warehouse HMI_pop_up_select_WIPs_select_wip_buttons{3}" : Push Button Data = PLC "HMI Data: Warehouse HMI".pop_up.select_WIPs.select_wip_buttons[3], 100 ms
   "HMI Data: Warehouse HMI_pop_up_select_WIPs_select_wip_buttons{4}" : Push Button Data = PLC "HMI Data: Warehouse HMI".pop_up.select_WIPs.select_wip_buttons[4], 100 ms
   "HMI Data: Warehouse HMI_pop_up_select_WIPs_select_wip_buttons{5}" : Push Button Data = PLC "HMI Data: Warehouse HMI".pop_up.select_WIPs.select_wip_buttons[5], 100 ms
   "HMI Data: Warehouse HMI_pop_up_select_WIPs_select_wip_buttons{6}" : Push Button Data = PLC "HMI Data: Warehouse HMI".pop_up.select_WIPs.select_wip_buttons[6], 100 ms
   "HMI Data: Warehouse HMI_pop_up_select_WIPs_close_screen" : Push Button Data = PLC "HMI Data: Warehouse HMI".pop_up.select_WIPs.close_screen, 100 ms
   "HMI Data: Warehouse HMI_pop_up_select_WIPs_nav_bar_hmi" : Nav Bar Data: HMI = PLC "HMI Data: Warehouse HMI".pop_up.select_WIPs.nav_bar.hmi, 100 ms

HMI tags "Part Call"
   "HMI Data: Warehouse HMI_partCall_row{0}" : Table Row = PLC "HMI Data: Warehouse HMI".partCall.row[0], 100 ms
   "HMI Data: Warehouse HMI_partCall_row{1}" : Table Row = PLC "HMI Data: Warehouse HMI".partCall.row[1], 100 ms
   "HMI Data: Warehouse HMI_partCall_row{10}" : Table Row = PLC "HMI Data: Warehouse HMI".partCall.row[10], 100 ms
   "HMI Data: Warehouse HMI_partCall_row{2}" : Table Row = PLC "HMI Data: Warehouse HMI".partCall.row[2], 100 ms
   "HMI Data: Warehouse HMI_partCall_row{3}" : Table Row = PLC "HMI Data: Warehouse HMI".partCall.row[3], 100 ms
   "HMI Data: Warehouse HMI_partCall_row{4}" : Table Row = PLC "HMI Data: Warehouse HMI".partCall.row[4], 100 ms
   "HMI Data: Warehouse HMI_partCall_row{5}" : Table Row = PLC "HMI Data: Warehouse HMI".partCall.row[5], 100 ms
   "HMI Data: Warehouse HMI_partCall_row{6}" : Table Row = PLC "HMI Data: Warehouse HMI".partCall.row[6], 100 ms
   "HMI Data: Warehouse HMI_partCall_row{7}" : Table Row = PLC "HMI Data: Warehouse HMI".partCall.row[7], 100 ms
   "HMI Data: Warehouse HMI_partCall_row{8}" : Table Row = PLC "HMI Data: Warehouse HMI".partCall.row[8], 100 ms
   "HMI Data: Warehouse HMI_partCall_row{9}" : Table Row = PLC "HMI Data: Warehouse HMI".partCall.row[9], 100 ms

